REGION Network 37: "flanco".niPul_MultiArr
   RUNG wire#powerrail
      N_Contact(operand := "iPul_MultiArr", bit := "xniPul_MultiArr")
      Coil( "flanco".niPul_MultiArr )
   END_RUNG
   // the same network as SCL:
   #_w1 := NOT "iPul_MultiArr" AND "xniPul_MultiArr";   // falling edge of "iPul_MultiArr"
   "xniPul_MultiArr" := "iPul_MultiArr";
   "flanco".niPul_MultiArr := #_w1;
END_REGION

REGION Network 38: "flanco".piPul_MultiAba
   RUNG wire#powerrail
      P_Contact(operand := "iPul_MultiAba", bit := "xpiPul_MultiAba")
      Coil( "flanco".piPul_MultiAba )
   END_RUNG
   // the same network as SCL:
   #_w1 := "iPul_MultiAba" AND NOT "xpiPul_MultiAba";   // rising edge of "iPul_MultiAba"
   "xpiPul_MultiAba" := "iPul_MultiAba";
   "flanco".piPul_MultiAba := #_w1;
END_REGION

REGION Network 39: "flanco".niPul_MultiAba
   RUNG wire#powerrail
      N_Contact(operand := "iPul_MultiAba", bit := "xniPul_MultiAba")
      Coil( "flanco".niPul_MultiAba )
   END_RUNG
   // the same network as SCL:
   #_w1 := NOT "iPul_MultiAba" AND "xniPul_MultiAba";   // falling edge of "iPul_MultiAba"
   "xniPul_MultiAba" := "iPul_MultiAba";
   "flanco".niPul_MultiAba := #_w1;
END_REGION

REGION Network 40: "flanco".piPul_MultiAde
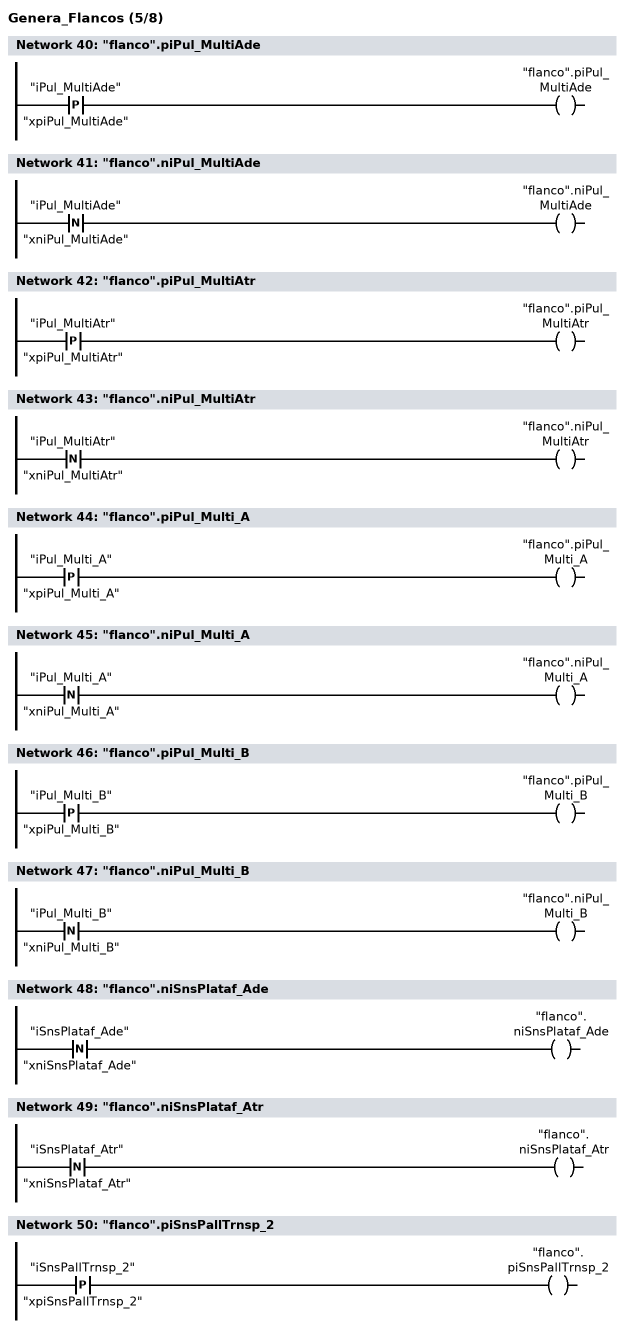
   RUNG wire#powerrail
      P_Contact(operand := "iPul_MultiAde", bit := "xpiPul_MultiAde")
      Coil( "flanco".piPul_MultiAde )
   END_RUNG
   // the same network as SCL:
   #_w1 := "iPul_MultiAde" AND NOT "xpiPul_MultiAde";   // rising edge of "iPul_MultiAde"
   "xpiPul_MultiAde" := "iPul_MultiAde";
   "flanco".piPul_MultiAde := #_w1;
END_REGION

REGION Network 41: "flanco".niPul_MultiAde
   RUNG wire#powerrail
      N_Contact(operand := "iPul_MultiAde", bit := "xniPul_MultiAde")
      Coil( "flanco".niPul_MultiAde )
   END_RUNG
   // the same network as SCL:
   #_w1 := NOT "iPul_MultiAde" AND "xniPul_MultiAde";   // falling edge of "iPul_MultiAde"
   "xniPul_MultiAde" := "iPul_MultiAde";
   "flanco".niPul_MultiAde := #_w1;
END_REGION

REGION Network 42: "flanco".piPul_MultiAtr
   RUNG wire#powerrail
      P_Contact(operand := "iPul_MultiAtr", bit := "xpiPul_MultiAtr")
      Coil( "flanco".piPul_MultiAtr )
   END_RUNG
   // the same network as SCL:
   #_w1 := "iPul_MultiAtr" AND NOT "xpiPul_MultiAtr";   // rising edge of "iPul_MultiAtr"
   "xpiPul_MultiAtr" := "iPul_MultiAtr";
   "flanco".piPul_MultiAtr := #_w1;
END_REGION

REGION Network 43: "flanco".niPul_MultiAtr
   RUNG wire#powerrail
      N_Contact(operand := "iPul_MultiAtr", bit := "xniPul_MultiAtr")
      Coil( "flanco".niPul_MultiAtr )
   END_RUNG
   // the same network as SCL:
   #_w1 := NOT "iPul_MultiAtr" AND "xniPul_MultiAtr";   // falling edge of "iPul_MultiAtr"
   "xniPul_MultiAtr" := "iPul_MultiAtr";
   "flanco".niPul_MultiAtr := #_w1;
END_REGION

REGION Network 44: "flanco".piPul_Multi_A
   RUNG wire#powerrail
      P_Contact(operand := "iPul_Multi_A", bit := "xpiPul_Multi_A")
      Coil( "flanco".piPul_Multi_A )
   END_RUNG
   // the same network as SCL:
   #_w1 := "iPul_Multi_A" AND NOT "xpiPul_Multi_A";   // rising edge of "iPul_Multi_A"
   "xpiPul_Multi_A" := "iPul_Multi_A";
   "flanco".piPul_Multi_A := #_w1;
END_REGION

REGION Network 45: "flanco".niPul_Multi_A
   RUNG wire#powerrail
      N_Contact(operand := "iPul_Multi_A", bit := "xniPul_Multi_A")
      Coil( "flanco".niPul_Multi_A )
   END_RUNG
   // the same network as SCL:
   #_w1 := NOT "iPul_Multi_A" AND "xniPul_Multi_A";   // falling edge of "iPul_Multi_A"
   "xniPul_Multi_A" := "iPul_Multi_A";
   "flanco".niPul_Multi_A := #_w1;
END_REGION

REGION Network 46: "flanco".piPul_Multi_B
   RUNG wire#powerrail
      P_Contact(operand := "iPul_Multi_B", bit := "xpiPul_Multi_B")
      Coil( "flanco".piPul_Multi_B )
   END_RUNG
   // the same network as SCL:
   #_w1 := "iPul_Multi_B" AND NOT "xpiPul_Multi_B";   // rising edge of "iPul_Multi_B"
   "xpiPul_Multi_B" := "iPul_Multi_B";
   "flanco".piPul_Multi_B := #_w1;
END_REGION

REGION Network 47: "flanco".niPul_Multi_B
   RUNG wire#powerrail
      N_Contact(operand := "iPul_Multi_B", bit := "xniPul_Multi_B")
      Coil( "flanco".niPul_Multi_B )
   END_RUNG
   // the same network as SCL:
   #_w1 := NOT "iPul_Multi_B" AND "xniPul_Multi_B";   // falling edge of "iPul_Multi_B"
   "xniPul_Multi_B" := "iPul_Multi_B";
   "flanco".niPul_Multi_B := #_w1;
END_REGION

REGION Network 48: "flanco".niSnsPlataf_Ade
   RUNG wire#powerrail
      N_Contact(operand := "iSnsPlataf_Ade", bit := "xniSnsPlataf_Ade")
      Coil( "flanco".niSnsPlataf_Ade )
   END_RUNG
   // the same network as SCL:
   #_w1 := NOT "iSnsPlataf_Ade" AND "xniSnsPlataf_Ade";   // falling edge of "iSnsPlataf_Ade"
   "xniSnsPlataf_Ade" := "iSnsPlataf_Ade";
   "flanco".niSnsPlataf_Ade := #_w1;
END_REGION

REGION Network 49: "flanco".niSnsPlataf_Atr
   RUNG wire#powerrail
      N_Contact(operand := "iSnsPlataf_Atr", bit := "xniSnsPlataf_Atr")
      Coil( "flanco".niSnsPlataf_Atr )
   END_RUNG
   // the same network as SCL:
   #_w1 := NOT "iSnsPlataf_Atr" AND "xniSnsPlataf_Atr";   // falling edge of "iSnsPlataf_Atr"
   "xniSnsPlataf_Atr" := "iSnsPlataf_Atr";
   "flanco".niSnsPlataf_Atr := #_w1;
END_REGION

REGION Network 50: "flanco".piSnsPallTrnsp_2
   RUNG wire#powerrail
      P_Contact(operand := "iSnsPallTrnsp_2", bit := "xpiSnsPallTrnsp_2")
      Coil( "flanco".piSnsPallTrnsp_2 )
   END_RUNG
   // the same network as SCL:
   #_w1 := "iSnsPallTrnsp_2" AND NOT "xpiSnsPallTrnsp_2";   // rising edge of "iSnsPallTrnsp_2"
   "xpiSnsPallTrnsp_2" := "iSnsPallTrnsp_2";
   "flanco".piSnsPallTrnsp_2 := #_w1;
END_REGION

REGION Network 51: "flanco".niSnsPallTrnsp_2
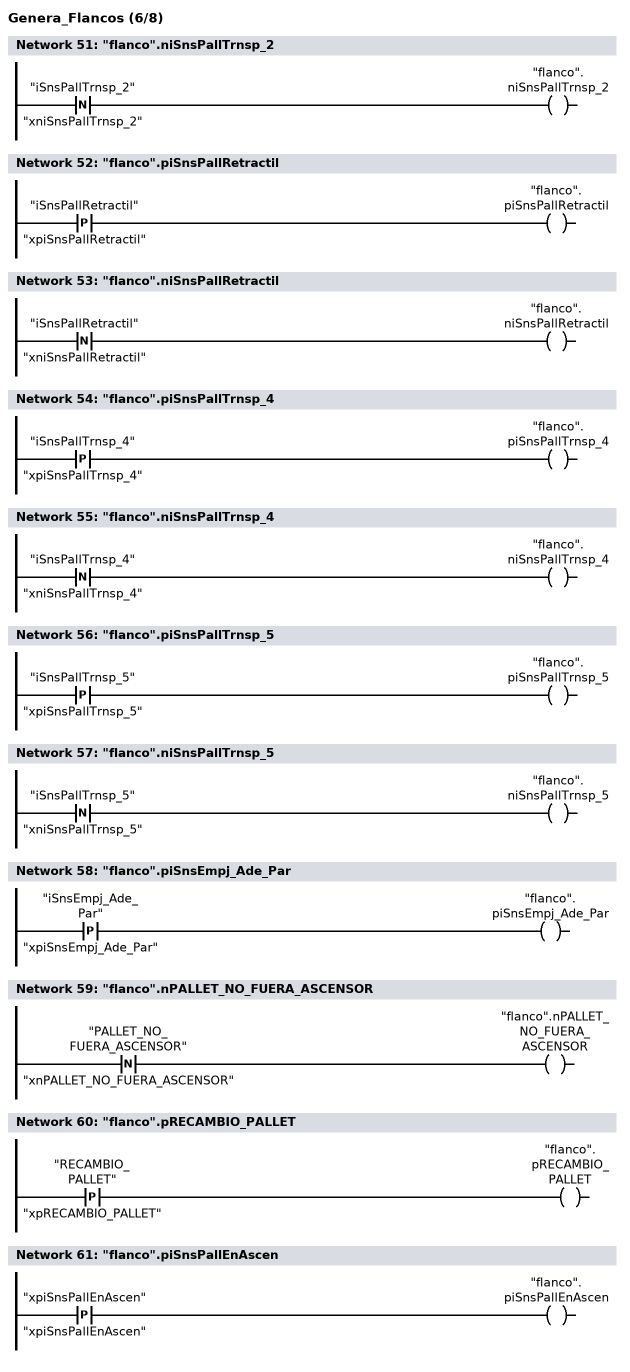
   RUNG wire#powerrail
      N_Contact(operand := "iSnsPallTrnsp_2", bit := "xniSnsPallTrnsp_2")
      Coil( "flanco".niSnsPallTrnsp_2 )
   END_RUNG
   // the same network as SCL:
   #_w1 := NOT "iSnsPallTrnsp_2" AND "xniSnsPallTrnsp_2";   // falling edge of "iSnsPallTrnsp_2"
   "xniSnsPallTrnsp_2" := "iSnsPallTrnsp_2";
   "flanco".niSnsPallTrnsp_2 := #_w1;
END_REGION

REGION Network 52: "flanco".piSnsPallRetractil
   RUNG wire#powerrail
      P_Contact(operand := "iSnsPallRetractil", bit := "xpiSnsPallRetractil")
      Coil( "flanco".piSnsPallRetractil )
   END_RUNG
   // the same network as SCL:
   #_w1 := "iSnsPallRetractil" AND NOT "xpiSnsPallRetractil";   // rising edge of "iSnsPallRetractil"
   "xpiSnsPallRetractil" := "iSnsPallRetractil";
   "flanco".piSnsPallRetractil := #_w1;
END_REGION

REGION Network 53: "flanco".niSnsPallRetractil
   RUNG wire#powerrail
      N_Contact(operand := "iSnsPallRetractil", bit := "xniSnsPallRetractil")
      Coil( "flanco".niSnsPallRetractil )
   END_RUNG
   // the same network as SCL:
   #_w1 := NOT "iSnsPallRetractil" AND "xniSnsPallRetractil";   // falling edge of "iSnsPallRetractil"
   "xniSnsPallRetractil" := "iSnsPallRetractil";
   "flanco".niSnsPallRetractil := #_w1;
END_REGION

REGION Network 54: "flanco".piSnsPallTrnsp_4
   RUNG wire#powerrail
      P_Contact(operand := "iSnsPallTrnsp_4", bit := "xpiSnsPallTrnsp_4")
      Coil( "flanco".piSnsPallTrnsp_4 )
   END_RUNG
   // the same network as SCL:
   #_w1 := "iSnsPallTrnsp_4" AND NOT "xpiSnsPallTrnsp_4";   // rising edge of "iSnsPallTrnsp_4"
   "xpiSnsPallTrnsp_4" := "iSnsPallTrnsp_4";
   "flanco".piSnsPallTrnsp_4 := #_w1;
END_REGION

REGION Network 55: "flanco".niSnsPallTrnsp_4
   RUNG wire#powerrail
      N_Contact(operand := "iSnsPallTrnsp_4", bit := "xniSnsPallTrnsp_4")
      Coil( "flanco".niSnsPallTrnsp_4 )
   END_RUNG
   // the same network as SCL:
   #_w1 := NOT "iSnsPallTrnsp_4" AND "xniSnsPallTrnsp_4";   // falling edge of "iSnsPallTrnsp_4"
   "xniSnsPallTrnsp_4" := "iSnsPallTrnsp_4";
   "flanco".niSnsPallTrnsp_4 := #_w1;
END_REGION

REGION Network 56: "flanco".piSnsPallTrnsp_5
   RUNG wire#powerrail
      P_Contact(operand := "iSnsPallTrnsp_5", bit := "xpiSnsPallTrnsp_5")
      Coil( "flanco".piSnsPallTrnsp_5 )
   END_RUNG
   // the same network as SCL:
   #_w1 := "iSnsPallTrnsp_5" AND NOT "xpiSnsPallTrnsp_5";   // rising edge of "iSnsPallTrnsp_5"
   "xpiSnsPallTrnsp_5" := "iSnsPallTrnsp_5";
   "flanco".piSnsPallTrnsp_5 := #_w1;
END_REGION

REGION Network 57: "flanco".niSnsPallTrnsp_5
   RUNG wire#powerrail
      N_Contact(operand := "iSnsPallTrnsp_5", bit := "xniSnsPallTrnsp_5")
      Coil( "flanco".niSnsPallTrnsp_5 )
   END_RUNG
   // the same network as SCL:
   #_w1 := NOT "iSnsPallTrnsp_5" AND "xniSnsPallTrnsp_5";   // falling edge of "iSnsPallTrnsp_5"
   "xniSnsPallTrnsp_5" := "iSnsPallTrnsp_5";
   "flanco".niSnsPallTrnsp_5 := #_w1;
END_REGION

REGION Network 58: "flanco".piSnsEmpj_Ade_Par
   RUNG wire#powerrail
      P_Contact(operand := "iSnsEmpj_Ade_Par", bit := "xpiSnsEmpj_Ade_Par")
      Coil( "flanco".piSnsEmpj_Ade_Par )
   END_RUNG
   // the same network as SCL:
   #_w1 := "iSnsEmpj_Ade_Par" AND NOT "xpiSnsEmpj_Ade_Par";   // rising edge of "iSnsEmpj_Ade_Par"
   "xpiSnsEmpj_Ade_Par" := "iSnsEmpj_Ade_Par";
   "flanco".piSnsEmpj_Ade_Par := #_w1;
END_REGION

REGION Network 59: "flanco".nPALLET_NO_FUERA_ASCENSOR
   RUNG wire#powerrail
      N_Contact(operand := "PALLET_NO_FUERA_ASCENSOR", bit := "xnPALLET_NO_FUERA_ASCENSOR")
      Coil( "flanco".nPALLET_NO_FUERA_ASCENSOR )
   END_RUNG
   // the same network as SCL:
   #_w1 := NOT "PALLET_NO_FUERA_ASCENSOR" AND "xnPALLET_NO_FUERA_ASCENSOR";   // falling edge of "PALLET_NO_FUERA_ASCENSOR"
   "xnPALLET_NO_FUERA_ASCENSOR" := "PALLET_NO_FUERA_ASCENSOR";
   "flanco".nPALLET_NO_FUERA_ASCENSOR := #_w1;
END_REGION

REGION Network 60: "flanco".pRECAMBIO_PALLET
   RUNG wire#powerrail
      P_Contact(operand := "RECAMBIO_PALLET", bit := "xpRECAMBIO_PALLET")
      Coil( "flanco".pRECAMBIO_PALLET )
   END_RUNG
   // the same network as SCL:
   #_w1 := "RECAMBIO_PALLET" AND NOT "xpRECAMBIO_PALLET";   // rising edge of "RECAMBIO_PALLET"
   "xpRECAMBIO_PALLET" := "RECAMBIO_PALLET";
   "flanco".pRECAMBIO_PALLET := #_w1;
END_REGION

REGION Network 61: "flanco".piSnsPallEnAscen
   RUNG wire#powerrail
      P_Contact(operand := "xpiSnsPallEnAscen", bit := "xpiSnsPallEnAscen")
      Coil( "flanco".piSnsPallEnAscen )
   END_RUNG
   // the same network as SCL:
   #_w1 := "xpiSnsPallEnAscen" AND NOT "xpiSnsPallEnAscen";   // rising edge of "xpiSnsPallEnAscen"
   "xpiSnsPallEnAscen" := "xpiSnsPallEnAscen";
   "flanco".piSnsPallEnAscen := #_w1;
END_REGION

REGION Network 62: "flanco".niSnsPallEnAscen
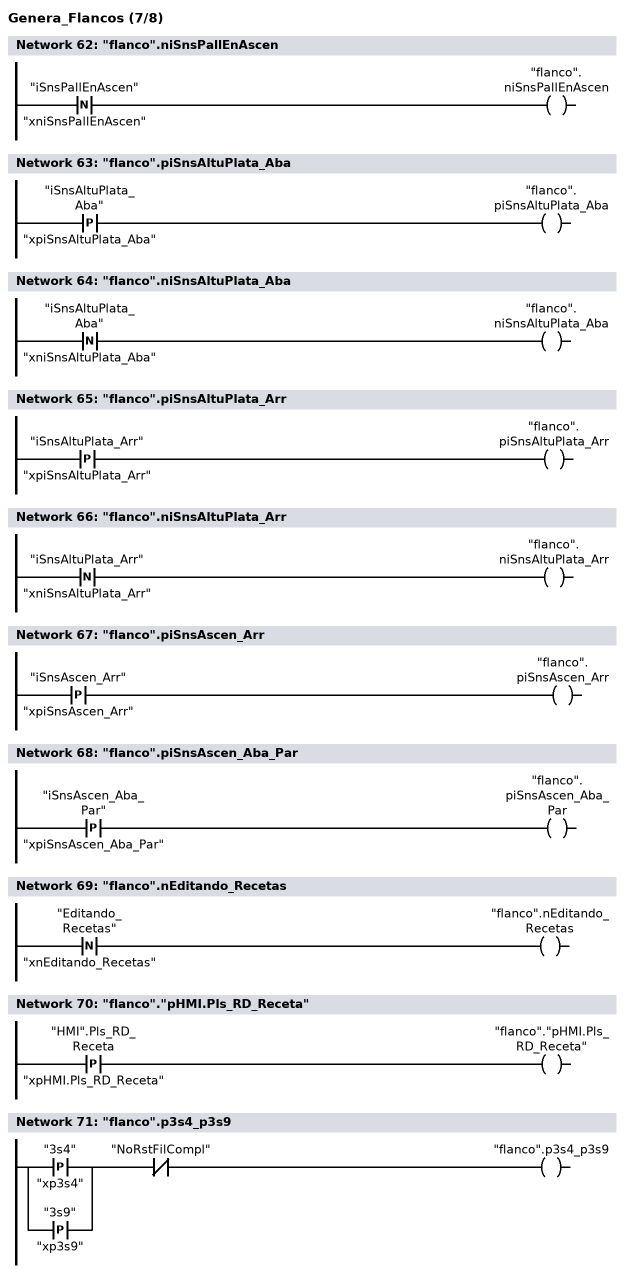
   RUNG wire#powerrail
      N_Contact(operand := "iSnsPallEnAscen", bit := "xniSnsPallEnAscen")
      Coil( "flanco".niSnsPallEnAscen )
   END_RUNG
   // the same network as SCL:
   #_w1 := NOT "iSnsPallEnAscen" AND "xniSnsPallEnAscen";   // falling edge of "iSnsPallEnAscen"
   "xniSnsPallEnAscen" := "iSnsPallEnAscen";
   "flanco".niSnsPallEnAscen := #_w1;
END_REGION

REGION Network 63: "flanco".piSnsAltuPlata_Aba
   RUNG wire#powerrail
      P_Contact(operand := "iSnsAltuPlata_Aba", bit := "xpiSnsAltuPlata_Aba")
      Coil( "flanco".piSnsAltuPlata_Aba )
   END_RUNG
   // the same network as SCL:
   #_w1 := "iSnsAltuPlata_Aba" AND NOT "xpiSnsAltuPlata_Aba";   // rising edge of "iSnsAltuPlata_Aba"
   "xpiSnsAltuPlata_Aba" := "iSnsAltuPlata_Aba";
   "flanco".piSnsAltuPlata_Aba := #_w1;
END_REGION

REGION Network 64: "flanco".niSnsAltuPlata_Aba
   RUNG wire#powerrail
      N_Contact(operand := "iSnsAltuPlata_Aba", bit := "xniSnsAltuPlata_Aba")
      Coil( "flanco".niSnsAltuPlata_Aba )
   END_RUNG
   // the same network as SCL:
   #_w1 := NOT "iSnsAltuPlata_Aba" AND "xniSnsAltuPlata_Aba";   // falling edge of "iSnsAltuPlata_Aba"
   "xniSnsAltuPlata_Aba" := "iSnsAltuPlata_Aba";
   "flanco".niSnsAltuPlata_Aba := #_w1;
END_REGION

REGION Network 65: "flanco".piSnsAltuPlata_Arr
   RUNG wire#powerrail
      P_Contact(operand := "iSnsAltuPlata_Arr", bit := "xpiSnsAltuPlata_Arr")
      Coil( "flanco".piSnsAltuPlata_Arr )
   END_RUNG
   // the same network as SCL:
   #_w1 := "iSnsAltuPlata_Arr" AND NOT "xpiSnsAltuPlata_Arr";   // rising edge of "iSnsAltuPlata_Arr"
   "xpiSnsAltuPlata_Arr" := "iSnsAltuPlata_Arr";
   "flanco".piSnsAltuPlata_Arr := #_w1;
END_REGION

REGION Network 66: "flanco".niSnsAltuPlata_Arr
   RUNG wire#powerrail
      N_Contact(operand := "iSnsAltuPlata_Arr", bit := "xniSnsAltuPlata_Arr")
      Coil( "flanco".niSnsAltuPlata_Arr )
   END_RUNG
   // the same network as SCL:
   #_w1 := NOT "iSnsAltuPlata_Arr" AND "xniSnsAltuPlata_Arr";   // falling edge of "iSnsAltuPlata_Arr"
   "xniSnsAltuPlata_Arr" := "iSnsAltuPlata_Arr";
   "flanco".niSnsAltuPlata_Arr := #_w1;
END_REGION

REGION Network 67: "flanco".piSnsAscen_Arr
   RUNG wire#powerrail
      P_Contact(operand := "iSnsAscen_Arr", bit := "xpiSnsAscen_Arr")
      Coil( "flanco".piSnsAscen_Arr )
   END_RUNG
   // the same network as SCL:
   #_w1 := "iSnsAscen_Arr" AND NOT "xpiSnsAscen_Arr";   // rising edge of "iSnsAscen_Arr"
   "xpiSnsAscen_Arr" := "iSnsAscen_Arr";
   "flanco".piSnsAscen_Arr := #_w1;
END_REGION

REGION Network 68: "flanco".piSnsAscen_Aba_Par
   RUNG wire#powerrail
      P_Contact(operand := "iSnsAscen_Aba_Par", bit := "xpiSnsAscen_Aba_Par")
      Coil( "flanco".piSnsAscen_Aba_Par )
   END_RUNG
   // the same network as SCL:
   #_w1 := "iSnsAscen_Aba_Par" AND NOT "xpiSnsAscen_Aba_Par";   // rising edge of "iSnsAscen_Aba_Par"
   "xpiSnsAscen_Aba_Par" := "iSnsAscen_Aba_Par";
   "flanco".piSnsAscen_Aba_Par := #_w1;
END_REGION

REGION Network 69: "flanco".nEditando_Recetas
   RUNG wire#powerrail
      N_Contact(operand := "Editando_Recetas", bit := "xnEditando_Recetas")
      Coil( "flanco".nEditando_Recetas )
   END_RUNG
   // the same network as SCL:
   #_w1 := NOT "Editando_Recetas" AND "xnEditando_Recetas";   // falling edge of "Editando_Recetas"
   "xnEditando_Recetas" := "Editando_Recetas";
   "flanco".nEditando_Recetas := #_w1;
END_REGION

REGION Network 70: "flanco"."pHMI.Pls_RD_Receta"
   RUNG wire#powerrail
      P_Contact(operand := "HMI".Pls_RD_Receta, bit := "xpHMI.Pls_RD_Receta")
      Coil( "flanco"."pHMI.Pls_RD_Receta" )
   END_RUNG
   // the same network as SCL:
   #_w1 := "HMI".Pls_RD_Receta AND NOT "xpHMI.Pls_RD_Receta";   // rising edge of "HMI".Pls_RD_Receta
   "xpHMI.Pls_RD_Receta" := "HMI".Pls_RD_Receta;
   "flanco"."pHMI.Pls_RD_Receta" := #_w1;
END_REGION

REGION Network 71: "flanco".p3s4_p3s9
   RUNG wire#powerrail
      P_Contact(operand := "3s4", bit := "xp3s4")
      wire#w1
      I_Contact( "NoRstFilCompl" )
      Coil( "flanco".p3s4_p3s9 )
   END_RUNG
   RUNG wire#powerrail
      P_Contact(operand := "3s9", bit := "xp3s9")
   END_RUNG wire#w1
   // the same network as SCL:
   #_w1 := "3s4" AND NOT "xp3s4";   // rising edge of "3s4"
   "xp3s4" := "3s4";
   #_w2 := "3s9" AND NOT "xp3s9";   // rising edge of "3s9"
   "xp3s9" := "3s9";
   "flanco".p3s4_p3s9 := (#_w1 OR #_w2) AND NOT "NoRstFilCompl";
END_REGION

REGION Network 72: "flanco"."pHMI.Pls_Inc_Figura_Sel"
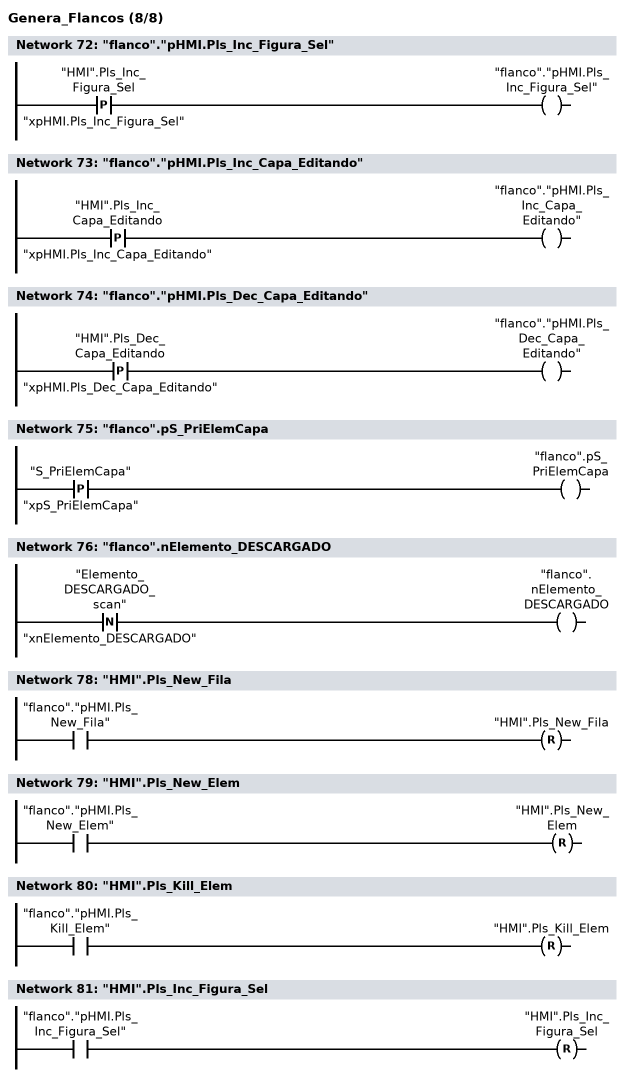
   RUNG wire#powerrail
      P_Contact(operand := "HMI".Pls_Inc_Figura_Sel, bit := "xpHMI.Pls_Inc_Figura_Sel")
      Coil( "flanco"."pHMI.Pls_Inc_Figura_Sel" )
   END_RUNG
   // the same network as SCL:
   #_w1 := "HMI".Pls_Inc_Figura_Sel AND NOT "xpHMI.Pls_Inc_Figura_Sel";   // rising edge of "HMI".Pls_Inc_Figura_Sel
   "xpHMI.Pls_Inc_Figura_Sel" := "HMI".Pls_Inc_Figura_Sel;
   "flanco"."pHMI.Pls_Inc_Figura_Sel" := #_w1;
END_REGION

REGION Network 73: "flanco"."pHMI.Pls_Inc_Capa_Editando"
   RUNG wire#powerrail
      P_Contact(operand := "HMI".Pls_Inc_Capa_Editando, bit := "xpHMI.Pls_Inc_Capa_Editando")
      Coil( "flanco"."pHMI.Pls_Inc_Capa_Editando" )
   END_RUNG
   // the same network as SCL:
   #_w1 := "HMI".Pls_Inc_Capa_Editando AND NOT "xpHMI.Pls_Inc_Capa_Editando";   // rising edge of "HMI".Pls_Inc_Capa_Editando
   "xpHMI.Pls_Inc_Capa_Editando" := "HMI".Pls_Inc_Capa_Editando;
   "flanco"."pHMI.Pls_Inc_Capa_Editando" := #_w1;
END_REGION

REGION Network 74: "flanco"."pHMI.Pls_Dec_Capa_Editando"
   RUNG wire#powerrail
      P_Contact(operand := "HMI".Pls_Dec_Capa_Editando, bit := "xpHMI.Pls_Dec_Capa_Editando")
      Coil( "flanco"."pHMI.Pls_Dec_Capa_Editando" )
   END_RUNG
   // the same network as SCL:
   #_w1 := "HMI".Pls_Dec_Capa_Editando AND NOT "xpHMI.Pls_Dec_Capa_Editando";   // rising edge of "HMI".Pls_Dec_Capa_Editando
   "xpHMI.Pls_Dec_Capa_Editando" := "HMI".Pls_Dec_Capa_Editando;
   "flanco"."pHMI.Pls_Dec_Capa_Editando" := #_w1;
END_REGION

REGION Network 75: "flanco".pS_PriElemCapa
   RUNG wire#powerrail
      P_Contact(operand := "S_PriElemCapa", bit := "xpS_PriElemCapa")
      Coil( "flanco".pS_PriElemCapa )
   END_RUNG
   // the same network as SCL:
   #_w1 := "S_PriElemCapa" AND NOT "xpS_PriElemCapa";   // rising edge of "S_PriElemCapa"
   "xpS_PriElemCapa" := "S_PriElemCapa";
   "flanco".pS_PriElemCapa := #_w1;
END_REGION

REGION Network 76: "flanco".nElemento_DESCARGADO
   RUNG wire#powerrail
      N_Contact(operand := "Elemento_DESCARGADO_scan", bit := "xnElemento_DESCARGADO")
      Coil( "flanco".nElemento_DESCARGADO )
   END_RUNG
   // the same network as SCL:
   #_w1 := NOT "Elemento_DESCARGADO_scan" AND "xnElemento_DESCARGADO";   // falling edge of "Elemento_DESCARGADO_scan"
   "xnElemento_DESCARGADO" := "Elemento_DESCARGADO_scan";
   "flanco".nElemento_DESCARGADO := #_w1;
END_REGION

REGION Network 77: ##################################################################
END_REGION

REGION Network 78: "HMI".Pls_New_Fila
   RUNG wire#powerrail
      Contact( "flanco"."pHMI.Pls_New_Fila" )
      R_Coil( "HMI".Pls_New_Fila )
   END_RUNG
   // the same network as SCL:
   IF "flanco"."pHMI.Pls_New_Fila" THEN "HMI".Pls_New_Fila := FALSE; END_IF;
END_REGION

REGION Network 79: "HMI".Pls_New_Elem
   RUNG wire#powerrail
      Contact( "flanco"."pHMI.Pls_New_Elem" )
      R_Coil( "HMI".Pls_New_Elem )
   END_RUNG
   // the same network as SCL:
   IF "flanco"."pHMI.Pls_New_Elem" THEN "HMI".Pls_New_Elem := FALSE; END_IF;
END_REGION

REGION Network 80: "HMI".Pls_Kill_Elem
   RUNG wire#powerrail
      Contact( "flanco"."pHMI.Pls_Kill_Elem" )
      R_Coil( "HMI".Pls_Kill_Elem )
   END_RUNG
   // the same network as SCL:
   IF "flanco"."pHMI.Pls_Kill_Elem" THEN "HMI".Pls_Kill_Elem := FALSE; END_IF;
END_REGION

REGION Network 81: "HMI".Pls_Inc_Figura_Sel
   RUNG wire#powerrail
      Contact( "flanco"."pHMI.Pls_Inc_Figura_Sel" )
      R_Coil( "HMI".Pls_Inc_Figura_Sel )
   END_RUNG
   // the same network as SCL:
   IF "flanco"."pHMI.Pls_Inc_Figura_Sel" THEN "HMI".Pls_Inc_Figura_Sel := FALSE; END_IF;
END_REGION
END_FUNCTION

FUNCTION "Cuenta_Cajas" : Void   // FC5, STL
{ S7_Optimized_Access := 'FALSE' }
VERSION : 0.1
BEGIN

REGION Network 1
         CLR;
         =     #Inc_1;
         =     #Inc_2;
         =     #Dec_1;
         =     #Dec_2;
         A     "S_ÚltFilCapa";
         A     "S_ÚltElemFila";
         =     #Ult_Elemento;
         ON    "S_PriElemCapa";
         O     "flanco".pS_PriElemCapa;
         =     #NoPri_Elemento;
END_REGION

REGION Network 2: Sumar Cajas
         L     "DB_Animación".Figura_SEL;
         L     2;
         <=I;
         JCN   AAAA;
   //    UN    #Ult_Elemento
         A     "Elemento_CARGADO";
         =     #Inc_1;
         JU    INCR;
   AAAA: TAK;
         L     3;
         ==I;
   //    UN    #Ult_Elemento
         A     "Elemento_CARGADO";
         =     #Inc_2;
   INCR: NOP   0;
END_REGION

REGION Network 3: Restar Cajas
         L     "DB_Animación".Figura_SEL;
         L     2;
         <=I;
         JCN   BBBB;
   //    U     #NoPri_Elemento
         A     "flanco".nElemento_DESCARGADO;
         =     #Dec_1;
         JU    DECR;
   BBBB: TAK;
         L     3;
         ==I;
   //    U     #NoPri_Elemento
         A     "flanco".nElemento_DESCARGADO;
         =     #Dec_2;
   DECR: NOP   0;
END_REGION

REGION Network 4: Cuenta las cajas en Empujador de Filas
         A     #Inc_1;  //Sumar de a una caja
         JCN   Mas1Caja;
         L     "Proceso Empujador".Cant_Cajas;
         L     DINT#1;
         +D;
         T     "Proceso Empujador".Cant_Cajas;
   Mas1Caja:NOP   0;
         A     #Inc_2;  //Sumar de a dos cajas
         JCN   Mas2Caja;
         L     "Proceso Empujador".Cant_Cajas;
         L     DINT#2;
         +D;
         T     "Proceso Empujador".Cant_Cajas;
   Mas2Caja:NOP   0;
         A     #Dec_1;  //Restar de a una caja
         JCN   Men1Caja;
         L     "Proceso Empujador".Cant_Cajas;
         L     DINT#1;
         -D;
         T     "Proceso Empujador".Cant_Cajas;
   Men1Caja:NOP   0;
         A     #Dec_2;  //Restar de a dos cajas
         JCN   Men2Caja;
         L     "Proceso Empujador".Cant_Cajas;
         L     DINT#2;
         -D;
         T     "Proceso Empujador".Cant_Cajas;
   Men2Caja:NOP   0;
         A     "HMI".Pls_ResetCajas;  //Resetear cajas producidas
         JCN   ReCaja;
         L     0;
         T     "Proceso Empujador".Cant_Cajas;
   ReCaja:NOP   0;
END_REGION
END_FUNCTION

FUNCTION "Genera_Señales" : Void   // FC16, LAD
{ S7_Optimized_Access := 'FALSE' }
VERSION : 0.1
BEGIN

REGION Network 1: ----------------------------------------------------------------- CARGA DE PALLETS -----------------------------------------------------------------¬
END_REGION

REGION Network 3: "Ascensor_Subir_Lento"
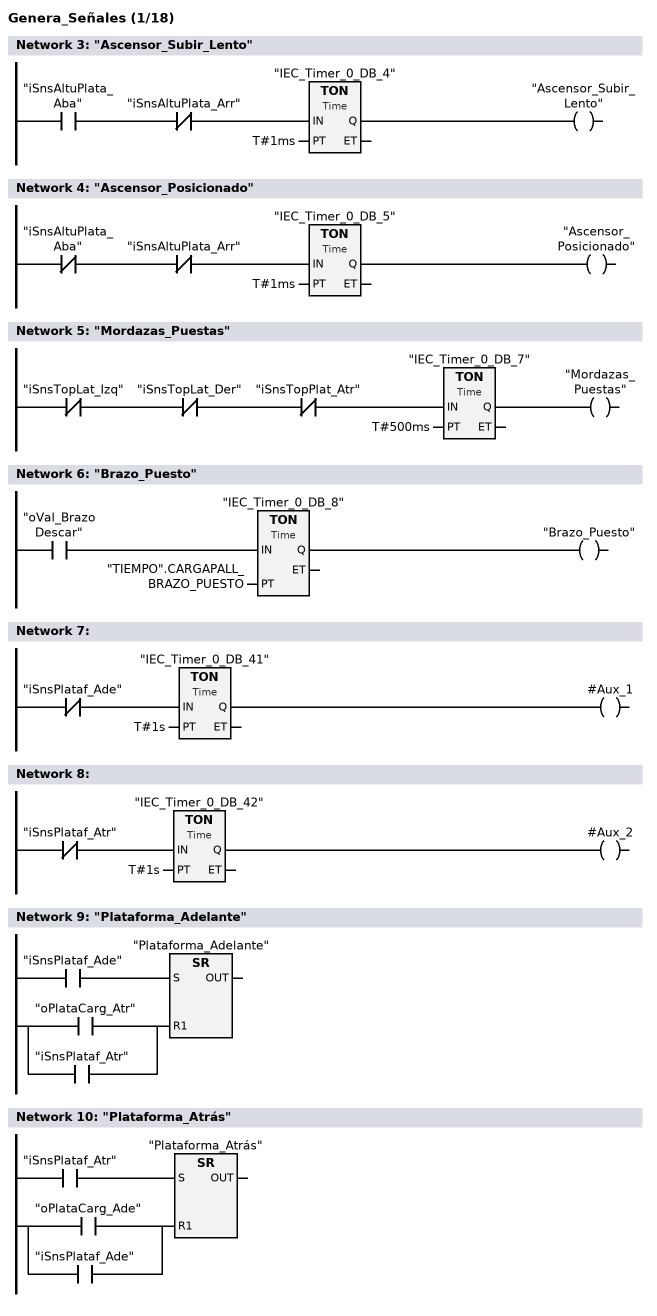
   "IEC_Timer_0_DB_4".TON(IN := "iSnsAltuPlata_Aba" AND NOT "iSnsAltuPlata_Arr", PT := T#1ms);
   "Ascensor_Subir_Lento" := "IEC_Timer_0_DB_4".Q;
END_REGION

REGION Network 4: "Ascensor_Posicionado"
   "IEC_Timer_0_DB_5".TON(IN := NOT "iSnsAltuPlata_Aba" AND NOT "iSnsAltuPlata_Arr", PT := T#1ms);
   "Ascensor_Posicionado" := "IEC_Timer_0_DB_5".Q;
END_REGION

REGION Network 5: "Mordazas_Puestas"
   "IEC_Timer_0_DB_7".TON(IN := NOT "iSnsTopLat_Izq" AND NOT "iSnsTopLat_Der" AND NOT "iSnsTopPlat_Atr",
                          PT := T#500ms);
   "Mordazas_Puestas" := "IEC_Timer_0_DB_7".Q;
END_REGION

REGION Network 6: "Brazo_Puesto"
   "IEC_Timer_0_DB_8".TON(IN := "oVal_BrazoDescar", PT := "TIEMPO".CARGAPALL_BRAZO_PUESTO);
   "Brazo_Puesto" := "IEC_Timer_0_DB_8".Q;
END_REGION

REGION Network 7
   "IEC_Timer_0_DB_41".TON(IN := NOT "iSnsPlataf_Ade", PT := T#1s);
   #Aux_1 := "IEC_Timer_0_DB_41".Q;
END_REGION

REGION Network 8
   "IEC_Timer_0_DB_42".TON(IN := NOT "iSnsPlataf_Atr", PT := T#1s);
   #Aux_2 := "IEC_Timer_0_DB_42".Q;
END_REGION

REGION Network 9: "Plataforma_Adelante"
   RUNG wire#powerrail
      Contact( "iSnsPlataf_Ade" )
      S_SR(operand := "Plataforma_Adelante", r1 := wire#w1)
   END_RUNG
   RUNG wire#powerrail
      Contact( "oPlataCarg_Atr" )
   END_RUNG wire#w1
   RUNG wire#powerrail
      Contact( "iSnsPlataf_Atr" )
   END_RUNG wire#w1
   // the same network as SCL:
   IF "iSnsPlataf_Ade" THEN
       "Plataforma_Adelante" := TRUE;   // SR flip-flop
   END_IF;
   IF "oPlataCarg_Atr" OR "iSnsPlataf_Atr" THEN "Plataforma_Adelante" := FALSE; END_IF;
END_REGION

REGION Network 10: "Plataforma_Atrás"
   RUNG wire#powerrail
      Contact( "iSnsPlataf_Atr" )
      S_SR(operand := "Plataforma_Atrás", r1 := wire#w1)
   END_RUNG
   RUNG wire#powerrail
      Contact( "oPlataCarg_Ade" )
   END_RUNG wire#w1
   RUNG wire#powerrail
      Contact( "iSnsPlataf_Ade" )
   END_RUNG wire#w1
   // the same network as SCL:
   IF "iSnsPlataf_Atr" THEN
       "Plataforma_Atrás" := TRUE;   // SR flip-flop
   END_IF;
   IF "oPlataCarg_Ade" OR "iSnsPlataf_Ade" THEN "Plataforma_Atrás" := FALSE; END_IF;
END_REGION

REGION Network 11: "PosiciónPlataf_Ade-Atr"
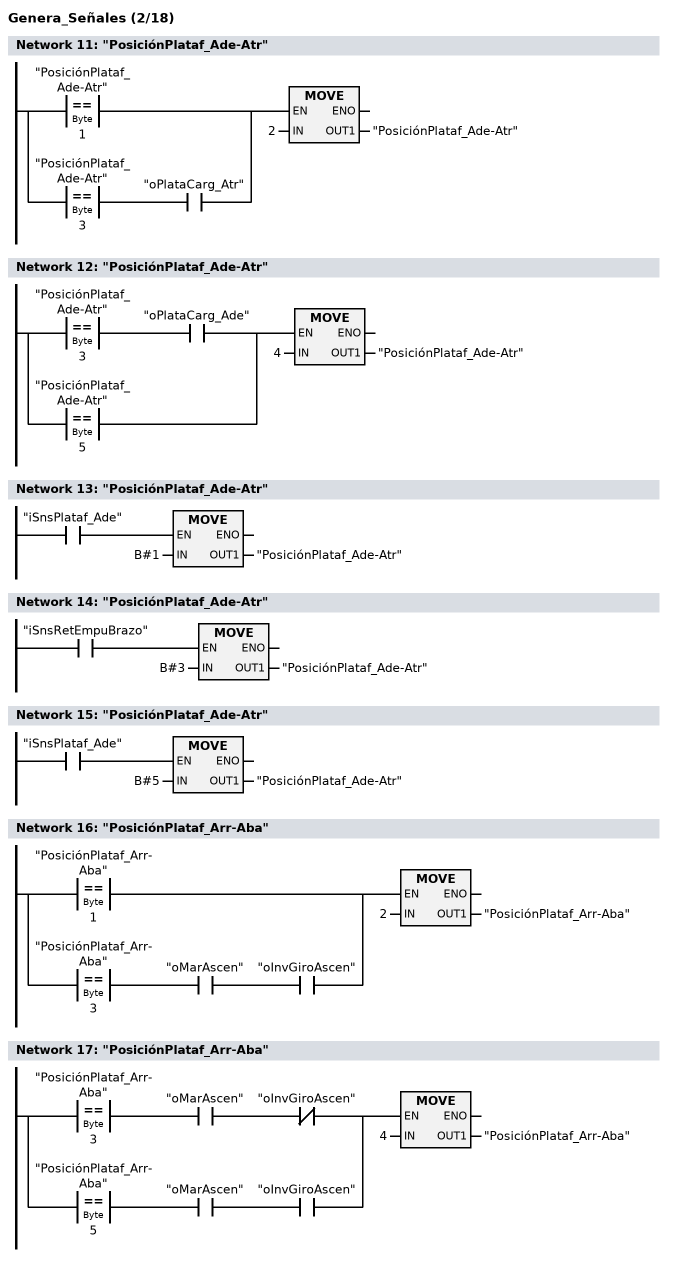
   RUNG wire#powerrail
      { S7_Templates := "SrcType := Byte" } EQ_Contact(in1 := "PosiciónPlataf_Ade-Atr", in2 := 1)
      wire#w1
      { S7_GenerateENO := "TRUE" } Move(in := 2, out1 => "PosiciónPlataf_Ade-Atr")
   END_RUNG
   RUNG wire#powerrail
      { S7_Templates := "SrcType := Byte" } EQ_Contact(in1 := "PosiciónPlataf_Ade-Atr", in2 := 3)
      Contact( "oPlataCarg_Atr" )
   END_RUNG wire#w1
   // the same network as SCL:
   IF ("PosiciónPlataf_Ade-Atr" = 1) OR (("PosiciónPlataf_Ade-Atr" = 3) AND "oPlataCarg_Atr") THEN
       "PosiciónPlataf_Ade-Atr" := 2;
   END_IF;
END_REGION

REGION Network 12: "PosiciónPlataf_Ade-Atr"
   RUNG wire#powerrail
      { S7_Templates := "SrcType := Byte" } EQ_Contact(in1 := "PosiciónPlataf_Ade-Atr", in2 := 3)
      Contact( "oPlataCarg_Ade" )
      wire#w1
      { S7_GenerateENO := "TRUE" } Move(in := 4, out1 => "PosiciónPlataf_Ade-Atr")
   END_RUNG
   RUNG wire#powerrail
      { S7_Templates := "SrcType := Byte" } EQ_Contact(in1 := "PosiciónPlataf_Ade-Atr", in2 := 5)
   END_RUNG wire#w1
   // the same network as SCL:
   IF (("PosiciónPlataf_Ade-Atr" = 3) AND "oPlataCarg_Ade") OR ("PosiciónPlataf_Ade-Atr" = 5) THEN
       "PosiciónPlataf_Ade-Atr" := 4;
   END_IF;
END_REGION

REGION Network 13: "PosiciónPlataf_Ade-Atr"
   RUNG wire#powerrail
      Contact( "iSnsPlataf_Ade" )
      { S7_GenerateENO := "TRUE" } Move(in := B#1, out1 => "PosiciónPlataf_Ade-Atr")
   END_RUNG
   // the same network as SCL:
   IF "iSnsPlataf_Ade" THEN "PosiciónPlataf_Ade-Atr" := B#1; END_IF;
END_REGION

REGION Network 14: "PosiciónPlataf_Ade-Atr"
   RUNG wire#powerrail
      Contact( "iSnsRetEmpuBrazo" )
      { S7_GenerateENO := "TRUE" } Move(in := B#3, out1 => "PosiciónPlataf_Ade-Atr")
   END_RUNG
   // the same network as SCL:
   IF "iSnsRetEmpuBrazo" THEN "PosiciónPlataf_Ade-Atr" := B#3; END_IF;
END_REGION

REGION Network 15: "PosiciónPlataf_Ade-Atr"
   RUNG wire#powerrail
      Contact( "iSnsPlataf_Ade" )
      { S7_GenerateENO := "TRUE" } Move(in := B#5, out1 => "PosiciónPlataf_Ade-Atr")
   END_RUNG
   // the same network as SCL:
   IF "iSnsPlataf_Ade" THEN "PosiciónPlataf_Ade-Atr" := B#5; END_IF;
END_REGION

REGION Network 16: "PosiciónPlataf_Arr-Aba"
   RUNG wire#powerrail
      { S7_Templates := "SrcType := Byte" } EQ_Contact(in1 := "PosiciónPlataf_Arr-Aba", in2 := 1)
      wire#w1
      { S7_GenerateENO := "TRUE" } Move(in := 2, out1 => "PosiciónPlataf_Arr-Aba")
   END_RUNG
   RUNG wire#powerrail
      { S7_Templates := "SrcType := Byte" } EQ_Contact(in1 := "PosiciónPlataf_Arr-Aba", in2 := 3)
      Contact( "oMarAscen" )
      Contact( "oInvGiroAscen" )
   END_RUNG wire#w1
   // the same network as SCL:
   IF ("PosiciónPlataf_Arr-Aba" = 1) OR (("PosiciónPlataf_Arr-Aba" = 3) AND "oMarAscen" AND "oInvGiroAscen") THEN
       "PosiciónPlataf_Arr-Aba" := 2;
   END_IF;
END_REGION

REGION Network 17: "PosiciónPlataf_Arr-Aba"
   RUNG wire#powerrail
      { S7_Templates := "SrcType := Byte" } EQ_Contact(in1 := "PosiciónPlataf_Arr-Aba", in2 := 3)
      Contact( "oMarAscen" )
      I_Contact( "oInvGiroAscen" )
      wire#w1
      { S7_GenerateENO := "TRUE" } Move(in := 4, out1 => "PosiciónPlataf_Arr-Aba")
   END_RUNG
   RUNG wire#powerrail
      { S7_Templates := "SrcType := Byte" } EQ_Contact(in1 := "PosiciónPlataf_Arr-Aba", in2 := 5)
      Contact( "oMarAscen" )
      Contact( "oInvGiroAscen" )
   END_RUNG wire#w1
   // the same network as SCL:
   IF (("PosiciónPlataf_Arr-Aba" = 3) AND "oMarAscen" AND NOT "oInvGiroAscen") OR (("PosiciónPlataf_Arr-Aba" = 5) AND "oMarAscen" AND "oInvGiroAscen") THEN
       "PosiciónPlataf_Arr-Aba" := 4;
   END_IF;
END_REGION

REGION Network 18: "PosiciónPlataf_Arr-Aba"